REGION Network 7: UN - Hold Command
   RUNG wire#powerrail
      Contact( "UN".PackML_Sts_Alarm.cmd_Hold )
      Contact( "UN".PackML_Sts_Alarm.moduleActive )
      wire#w1
      Coil( "UN".PackML_Sts.cmd_Hold )
   END_RUNG
   RUNG wire#powerrail
      Contact( "EM00".PackML_Sts.Unit.cmd_Hold )
      Contact( "EM00".PackML_Sts.Unit.moduleActive )
   END_RUNG wire#w1
   RUNG wire#powerrail
      Contact( "EM01".PackML_Sts.Unit.cmd_Hold )
      Contact( "EM01".PackML_Sts.Unit.moduleActive )
   END_RUNG wire#w1
   RUNG wire#powerrail
      Contact( "EM02".PackML_Sts.Unit.cmd_Hold )
      Contact( "EM02".PackML_Sts.Unit.moduleActive )
   END_RUNG wire#w1
   // the same network as SCL:
   "UN".PackML_Sts.cmd_Hold := ("UN".PackML_Sts_Alarm.cmd_Hold AND "UN".PackML_Sts_Alarm.moduleActive) OR ("EM00".PackML_Sts.Unit.cmd_Hold AND "EM00".PackML_Sts.Unit.moduleActive) OR ("EM01".PackML_Sts.Unit.cmd_Hold AND "EM01".PackML_Sts.Unit.moduleActive) OR ("EM02".PackML_Sts.Unit.cmd_Hold AND "EM02".PackML_Sts.Unit.moduleActive);
END_REGION

REGION Network 8: UN - Holding State Complete
   RUNG wire#powerrail
      Contact( "UN".PackML_Sts_Alarm.sts_Holding_SC )
      wire#w1
      Contact( "EM00".PackML_Sts.Unit.sts_Holding_SC )
      wire#w2
      Contact( "EM01".PackML_Sts.Unit.sts_Holding_SC )
      wire#w3
      Contact( "EM02".PackML_Sts.Unit.sts_Holding_SC )
      wire#w4
      Coil( "UN".PackML_Sts.sts_Holding_SC )
   END_RUNG
   RUNG wire#powerrail
      I_Contact( "UN".PackML_Sts_Alarm.moduleActive )
   END_RUNG wire#w1
   RUNG wire#w1
      I_Contact( "EM00".PackML_Sts.Unit.moduleActive )
   END_RUNG wire#w2
   RUNG wire#w2
      I_Contact( "EM01".PackML_Sts.Unit.moduleActive )
   END_RUNG wire#w3
   RUNG wire#w3
      I_Contact( "EM02".PackML_Sts.Unit.moduleActive )
   END_RUNG wire#w4
   // the same network as SCL:
   "UN".PackML_Sts.sts_Holding_SC := ("UN".PackML_Sts_Alarm.sts_Holding_SC OR NOT "UN".PackML_Sts_Alarm.moduleActive) AND ("EM00".PackML_Sts.Unit.sts_Holding_SC OR NOT "EM00".PackML_Sts.Unit.moduleActive) AND ("EM01".PackML_Sts.Unit.sts_Holding_SC OR NOT "EM01".PackML_Sts.Unit.moduleActive) AND ("EM02".PackML_Sts.Unit.sts_Holding_SC OR NOT "EM02".PackML_Sts.Unit.moduleActive);
END_REGION

REGION Network 9: UN - UnHold Command
   RUNG wire#powerrail
      Contact( "UN".PackML_Sts_Alarm.cmd_UnHold )
      wire#w1
      Contact( "EM00".PackML_Sts.Unit.cmd_UnHold )
      wire#w2
      Contact( "EM01".PackML_Sts.Unit.cmd_UnHold )
      wire#w3
      Contact( "EM02".PackML_Sts.Unit.cmd_UnHold )
      wire#w4
      Coil( "UN".PackML_Sts.cmd_UnHold )
   END_RUNG
   RUNG wire#powerrail
      I_Contact( "UN".PackML_Sts_Alarm.moduleActive )
   END_RUNG wire#w1
   RUNG wire#w1
      I_Contact( "EM00".PackML_Sts.Unit.moduleActive )
   END_RUNG wire#w2
   RUNG wire#w2
      I_Contact( "EM01".PackML_Sts.Unit.moduleActive )
   END_RUNG wire#w3
   RUNG wire#w3
      I_Contact( "EM02".PackML_Sts.Unit.moduleActive )
   END_RUNG wire#w4
   // the same network as SCL:
   "UN".PackML_Sts.cmd_UnHold := ("UN".PackML_Sts_Alarm.cmd_UnHold OR NOT "UN".PackML_Sts_Alarm.moduleActive) AND ("EM00".PackML_Sts.Unit.cmd_UnHold OR NOT "EM00".PackML_Sts.Unit.moduleActive) AND ("EM01".PackML_Sts.Unit.cmd_UnHold OR NOT "EM01".PackML_Sts.Unit.moduleActive) AND ("EM02".PackML_Sts.Unit.cmd_UnHold OR NOT "EM02".PackML_Sts.Unit.moduleActive);
END_REGION

REGION Network 10: UN - UnHolding State Complete
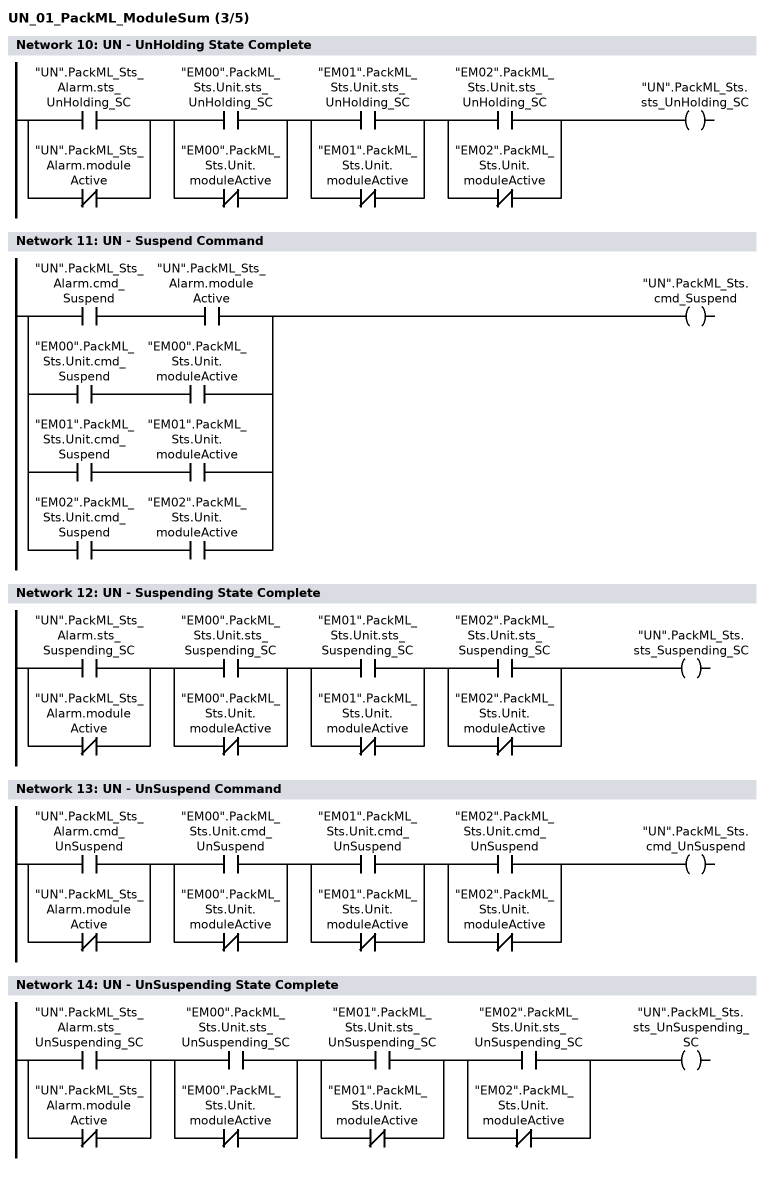
   RUNG wire#powerrail
      Contact( "UN".PackML_Sts_Alarm.sts_UnHolding_SC )
      wire#w1
      Contact( "EM00".PackML_Sts.Unit.sts_UnHolding_SC )
      wire#w2
      Contact( "EM01".PackML_Sts.Unit.sts_UnHolding_SC )
      wire#w3
      Contact( "EM02".PackML_Sts.Unit.sts_UnHolding_SC )
      wire#w4
      Coil( "UN".PackML_Sts.sts_UnHolding_SC )
   END_RUNG
   RUNG wire#powerrail
      I_Contact( "UN".PackML_Sts_Alarm.moduleActive )
   END_RUNG wire#w1
   RUNG wire#w1
      I_Contact( "EM00".PackML_Sts.Unit.moduleActive )
   END_RUNG wire#w2
   RUNG wire#w2
      I_Contact( "EM01".PackML_Sts.Unit.moduleActive )
   END_RUNG wire#w3
   RUNG wire#w3
      I_Contact( "EM02".PackML_Sts.Unit.moduleActive )
   END_RUNG wire#w4
   // the same network as SCL:
   "UN".PackML_Sts.sts_UnHolding_SC := ("UN".PackML_Sts_Alarm.sts_UnHolding_SC OR NOT "UN".PackML_Sts_Alarm.moduleActive) AND ("EM00".PackML_Sts.Unit.sts_UnHolding_SC OR NOT "EM00".PackML_Sts.Unit.moduleActive) AND ("EM01".PackML_Sts.Unit.sts_UnHolding_SC OR NOT "EM01".PackML_Sts.Unit.moduleActive) AND ("EM02".PackML_Sts.Unit.sts_UnHolding_SC OR NOT "EM02".PackML_Sts.Unit.moduleActive);
END_REGION

REGION Network 11: UN - Suspend Command
   RUNG wire#powerrail
      Contact( "UN".PackML_Sts_Alarm.cmd_Suspend )
      Contact( "UN".PackML_Sts_Alarm.moduleActive )
      wire#w1
      Coil( "UN".PackML_Sts.cmd_Suspend )
   END_RUNG
   RUNG wire#powerrail
      Contact( "EM00".PackML_Sts.Unit.cmd_Suspend )
      Contact( "EM00".PackML_Sts.Unit.moduleActive )
   END_RUNG wire#w1
   RUNG wire#powerrail
      Contact( "EM01".PackML_Sts.Unit.cmd_Suspend )
      Contact( "EM01".PackML_Sts.Unit.moduleActive )
   END_RUNG wire#w1
   RUNG wire#powerrail
      Contact( "EM02".PackML_Sts.Unit.cmd_Suspend )
      Contact( "EM02".PackML_Sts.Unit.moduleActive )
   END_RUNG wire#w1
   // the same network as SCL:
   "UN".PackML_Sts.cmd_Suspend := ("UN".PackML_Sts_Alarm.cmd_Suspend AND "UN".PackML_Sts_Alarm.moduleActive) OR ("EM00".PackML_Sts.Unit.cmd_Suspend AND "EM00".PackML_Sts.Unit.moduleActive) OR ("EM01".PackML_Sts.Unit.cmd_Suspend AND "EM01".PackML_Sts.Unit.moduleActive) OR ("EM02".PackML_Sts.Unit.cmd_Suspend AND "EM02".PackML_Sts.Unit.moduleActive);
END_REGION

REGION Network 12: UN - Suspending State Complete
   RUNG wire#powerrail
      Contact( "UN".PackML_Sts_Alarm.sts_Suspending_SC )
      wire#w1
      Contact( "EM00".PackML_Sts.Unit.sts_Suspending_SC )
      wire#w2
      Contact( "EM01".PackML_Sts.Unit.sts_Suspending_SC )
      wire#w3
      Contact( "EM02".PackML_Sts.Unit.sts_Suspending_SC )
      wire#w4
      Coil( "UN".PackML_Sts.sts_Suspending_SC )
   END_RUNG
   RUNG wire#powerrail
      I_Contact( "UN".PackML_Sts_Alarm.moduleActive )
   END_RUNG wire#w1
   RUNG wire#w1
      I_Contact( "EM00".PackML_Sts.Unit.moduleActive )
   END_RUNG wire#w2
   RUNG wire#w2
      I_Contact( "EM01".PackML_Sts.Unit.moduleActive )
   END_RUNG wire#w3
   RUNG wire#w3
      I_Contact( "EM02".PackML_Sts.Unit.moduleActive )
   END_RUNG wire#w4
   // the same network as SCL:
   "UN".PackML_Sts.sts_Suspending_SC := ("UN".PackML_Sts_Alarm.sts_Suspending_SC OR NOT "UN".PackML_Sts_Alarm.moduleActive) AND ("EM00".PackML_Sts.Unit.sts_Suspending_SC OR NOT "EM00".PackML_Sts.Unit.moduleActive) AND ("EM01".PackML_Sts.Unit.sts_Suspending_SC OR NOT "EM01".PackML_Sts.Unit.moduleActive) AND ("EM02".PackML_Sts.Unit.sts_Suspending_SC OR NOT "EM02".PackML_Sts.Unit.moduleActive);
END_REGION

REGION Network 13: UN - UnSuspend Command
   RUNG wire#powerrail
      Contact( "UN".PackML_Sts_Alarm.cmd_UnSuspend )
      wire#w1
      Contact( "EM00".PackML_Sts.Unit.cmd_UnSuspend )
      wire#w2
      Contact( "EM01".PackML_Sts.Unit.cmd_UnSuspend )
      wire#w3
      Contact( "EM02".PackML_Sts.Unit.cmd_UnSuspend )
      wire#w4
      Coil( "UN".PackML_Sts.cmd_UnSuspend )
   END_RUNG
   RUNG wire#powerrail
      I_Contact( "UN".PackML_Sts_Alarm.moduleActive )
   END_RUNG wire#w1
   RUNG wire#w1
      I_Contact( "EM00".PackML_Sts.Unit.moduleActive )
   END_RUNG wire#w2
   RUNG wire#w2
      I_Contact( "EM01".PackML_Sts.Unit.moduleActive )
   END_RUNG wire#w3
   RUNG wire#w3
      I_Contact( "EM02".PackML_Sts.Unit.moduleActive )
   END_RUNG wire#w4
   // the same network as SCL:
   "UN".PackML_Sts.cmd_UnSuspend := ("UN".PackML_Sts_Alarm.cmd_UnSuspend OR NOT "UN".PackML_Sts_Alarm.moduleActive) AND ("EM00".PackML_Sts.Unit.cmd_UnSuspend OR NOT "EM00".PackML_Sts.Unit.moduleActive) AND ("EM01".PackML_Sts.Unit.cmd_UnSuspend OR NOT "EM01".PackML_Sts.Unit.moduleActive) AND ("EM02".PackML_Sts.Unit.cmd_UnSuspend OR NOT "EM02".PackML_Sts.Unit.moduleActive);
END_REGION

REGION Network 14: UN - UnSuspending State Complete
   RUNG wire#powerrail
      Contact( "UN".PackML_Sts_Alarm.sts_UnSuspending_SC )
      wire#w1
      Contact( "EM00".PackML_Sts.Unit.sts_UnSuspending_SC )
      wire#w2
      Contact( "EM01".PackML_Sts.Unit.sts_UnSuspending_SC )
      wire#w3
      Contact( "EM02".PackML_Sts.Unit.sts_UnSuspending_SC )
      wire#w4
      Coil( "UN".PackML_Sts.sts_UnSuspending_SC )
   END_RUNG
   RUNG wire#powerrail
      I_Contact( "UN".PackML_Sts_Alarm.moduleActive )
   END_RUNG wire#w1
   RUNG wire#w1
      I_Contact( "EM00".PackML_Sts.Unit.moduleActive )
   END_RUNG wire#w2
   RUNG wire#w2
      I_Contact( "EM01".PackML_Sts.Unit.moduleActive )
   END_RUNG wire#w3
   RUNG wire#w3
      I_Contact( "EM02".PackML_Sts.Unit.moduleActive )
   END_RUNG wire#w4
   // the same network as SCL:
   "UN".PackML_Sts.sts_UnSuspending_SC := ("UN".PackML_Sts_Alarm.sts_UnSuspending_SC OR NOT "UN".PackML_Sts_Alarm.moduleActive) AND ("EM00".PackML_Sts.Unit.sts_UnSuspending_SC OR NOT "EM00".PackML_Sts.Unit.moduleActive) AND ("EM01".PackML_Sts.Unit.sts_UnSuspending_SC OR NOT "EM01".PackML_Sts.Unit.moduleActive) AND ("EM02".PackML_Sts.Unit.sts_UnSuspending_SC OR NOT "EM02".PackML_Sts.Unit.moduleActive);
END_REGION

REGION Network 15: UN - Abort Command
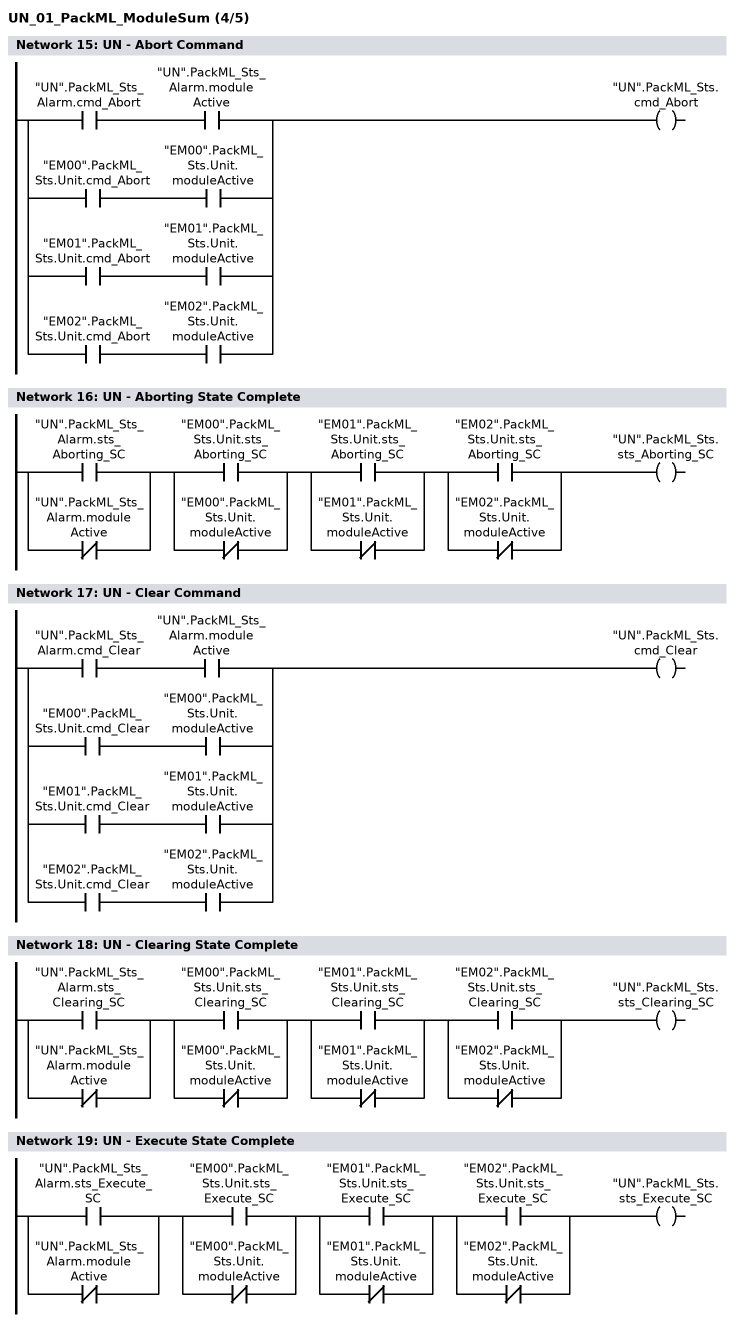
   RUNG wire#powerrail
      Contact( "UN".PackML_Sts_Alarm.cmd_Abort )
      Contact( "UN".PackML_Sts_Alarm.moduleActive )
      wire#w1
      Coil( "UN".PackML_Sts.cmd_Abort )
   END_RUNG
   RUNG wire#powerrail
      Contact( "EM00".PackML_Sts.Unit.cmd_Abort )
      Contact( "EM00".PackML_Sts.Unit.moduleActive )
   END_RUNG wire#w1
   RUNG wire#powerrail
      Contact( "EM01".PackML_Sts.Unit.cmd_Abort )
      Contact( "EM01".PackML_Sts.Unit.moduleActive )
   END_RUNG wire#w1
   RUNG wire#powerrail
      Contact( "EM02".PackML_Sts.Unit.cmd_Abort )
      Contact( "EM02".PackML_Sts.Unit.moduleActive )
   END_RUNG wire#w1
   // the same network as SCL:
   "UN".PackML_Sts.cmd_Abort := ("UN".PackML_Sts_Alarm.cmd_Abort AND "UN".PackML_Sts_Alarm.moduleActive) OR ("EM00".PackML_Sts.Unit.cmd_Abort AND "EM00".PackML_Sts.Unit.moduleActive) OR ("EM01".PackML_Sts.Unit.cmd_Abort AND "EM01".PackML_Sts.Unit.moduleActive) OR ("EM02".PackML_Sts.Unit.cmd_Abort AND "EM02".PackML_Sts.Unit.moduleActive);
END_REGION

REGION Network 16: UN - Aborting State Complete
   RUNG wire#powerrail
      Contact( "UN".PackML_Sts_Alarm.sts_Aborting_SC )
      wire#w1
      Contact( "EM00".PackML_Sts.Unit.sts_Aborting_SC )
      wire#w2
      Contact( "EM01".PackML_Sts.Unit.sts_Aborting_SC )
      wire#w3
      Contact( "EM02".PackML_Sts.Unit.sts_Aborting_SC )
      wire#w4
      Coil( "UN".PackML_Sts.sts_Aborting_SC )
   END_RUNG
   RUNG wire#powerrail
      I_Contact( "UN".PackML_Sts_Alarm.moduleActive )
   END_RUNG wire#w1
   RUNG wire#w1
      I_Contact( "EM00".PackML_Sts.Unit.moduleActive )
   END_RUNG wire#w2
   RUNG wire#w2
      I_Contact( "EM01".PackML_Sts.Unit.moduleActive )
   END_RUNG wire#w3
   RUNG wire#w3
      I_Contact( "EM02".PackML_Sts.Unit.moduleActive )
   END_RUNG wire#w4
   // the same network as SCL:
   "UN".PackML_Sts.sts_Aborting_SC := ("UN".PackML_Sts_Alarm.sts_Aborting_SC OR NOT "UN".PackML_Sts_Alarm.moduleActive) AND ("EM00".PackML_Sts.Unit.sts_Aborting_SC OR NOT "EM00".PackML_Sts.Unit.moduleActive) AND ("EM01".PackML_Sts.Unit.sts_Aborting_SC OR NOT "EM01".PackML_Sts.Unit.moduleActive) AND ("EM02".PackML_Sts.Unit.sts_Aborting_SC OR NOT "EM02".PackML_Sts.Unit.moduleActive);
END_REGION

REGION Network 17: UN - Clear Command
   RUNG wire#powerrail
      Contact( "UN".PackML_Sts_Alarm.cmd_Clear )
      Contact( "UN".PackML_Sts_Alarm.moduleActive )
      wire#w1
      Coil( "UN".PackML_Sts.cmd_Clear )
   END_RUNG
   RUNG wire#powerrail
      Contact( "EM00".PackML_Sts.Unit.cmd_Clear )
      Contact( "EM00".PackML_Sts.Unit.moduleActive )
   END_RUNG wire#w1
   RUNG wire#powerrail
      Contact( "EM01".PackML_Sts.Unit.cmd_Clear )
      Contact( "EM01".PackML_Sts.Unit.moduleActive )
   END_RUNG wire#w1
   RUNG wire#powerrail
      Contact( "EM02".PackML_Sts.Unit.cmd_Clear )
      Contact( "EM02".PackML_Sts.Unit.moduleActive )
   END_RUNG wire#w1
   // the same network as SCL:
   "UN".PackML_Sts.cmd_Clear := ("UN".PackML_Sts_Alarm.cmd_Clear AND "UN".PackML_Sts_Alarm.moduleActive) OR ("EM00".PackML_Sts.Unit.cmd_Clear AND "EM00".PackML_Sts.Unit.moduleActive) OR ("EM01".PackML_Sts.Unit.cmd_Clear AND "EM01".PackML_Sts.Unit.moduleActive) OR ("EM02".PackML_Sts.Unit.cmd_Clear AND "EM02".PackML_Sts.Unit.moduleActive);
END_REGION

REGION Network 18: UN - Clearing State Complete
   RUNG wire#powerrail
      Contact( "UN".PackML_Sts_Alarm.sts_Clearing_SC )
      wire#w1
      Contact( "EM00".PackML_Sts.Unit.sts_Clearing_SC )
      wire#w2
      Contact( "EM01".PackML_Sts.Unit.sts_Clearing_SC )
      wire#w3
      Contact( "EM02".PackML_Sts.Unit.sts_Clearing_SC )
      wire#w4
      Coil( "UN".PackML_Sts.sts_Clearing_SC )
   END_RUNG
   RUNG wire#powerrail
      I_Contact( "UN".PackML_Sts_Alarm.moduleActive )
   END_RUNG wire#w1
   RUNG wire#w1
      I_Contact( "EM00".PackML_Sts.Unit.moduleActive )
   END_RUNG wire#w2
   RUNG wire#w2
      I_Contact( "EM01".PackML_Sts.Unit.moduleActive )
   END_RUNG wire#w3
   RUNG wire#w3
      I_Contact( "EM02".PackML_Sts.Unit.moduleActive )
   END_RUNG wire#w4
   // the same network as SCL:
   "UN".PackML_Sts.sts_Clearing_SC := ("UN".PackML_Sts_Alarm.sts_Clearing_SC OR NOT "UN".PackML_Sts_Alarm.moduleActive) AND ("EM00".PackML_Sts.Unit.sts_Clearing_SC OR NOT "EM00".PackML_Sts.Unit.moduleActive) AND ("EM01".PackML_Sts.Unit.sts_Clearing_SC OR NOT "EM01".PackML_Sts.Unit.moduleActive) AND ("EM02".PackML_Sts.Unit.sts_Clearing_SC OR NOT "EM02".PackML_Sts.Unit.moduleActive);
END_REGION

REGION Network 19: UN - Execute State Complete
   RUNG wire#powerrail
      Contact( "UN".PackML_Sts_Alarm.sts_Execute_SC )
      wire#w1
      Contact( "EM00".PackML_Sts.Unit.sts_Execute_SC )
      wire#w2
      Contact( "EM01".PackML_Sts.Unit.sts_Execute_SC )
      wire#w3
      Contact( "EM02".PackML_Sts.Unit.sts_Execute_SC )
      wire#w4
      Coil( "UN".PackML_Sts.sts_Execute_SC )
   END_RUNG
   RUNG wire#powerrail
      I_Contact( "UN".PackML_Sts_Alarm.moduleActive )
   END_RUNG wire#w1
   RUNG wire#w1
      I_Contact( "EM00".PackML_Sts.Unit.moduleActive )
   END_RUNG wire#w2
   RUNG wire#w2
      I_Contact( "EM01".PackML_Sts.Unit.moduleActive )
   END_RUNG wire#w3
   RUNG wire#w3
      I_Contact( "EM02".PackML_Sts.Unit.moduleActive )
   END_RUNG wire#w4
   // the same network as SCL:
   "UN".PackML_Sts.sts_Execute_SC := ("UN".PackML_Sts_Alarm.sts_Execute_SC OR NOT "UN".PackML_Sts_Alarm.moduleActive) AND ("EM00".PackML_Sts.Unit.sts_Execute_SC OR NOT "EM00".PackML_Sts.Unit.moduleActive) AND ("EM01".PackML_Sts.Unit.sts_Execute_SC OR NOT "EM01".PackML_Sts.Unit.moduleActive) AND ("EM02".PackML_Sts.Unit.sts_Execute_SC OR NOT "EM02".PackML_Sts.Unit.moduleActive);
END_REGION

REGION Network 20: UN - Completing State Complete
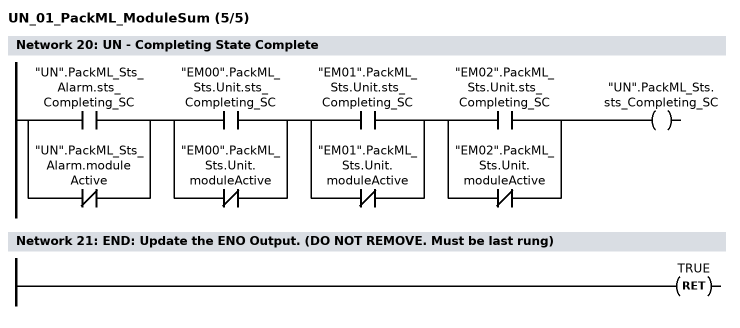
   RUNG wire#powerrail
      Contact( "UN".PackML_Sts_Alarm.sts_Completing_SC )
      wire#w1
      Contact( "EM00".PackML_Sts.Unit.sts_Completing_SC )
      wire#w2
      Contact( "EM01".PackML_Sts.Unit.sts_Completing_SC )
      wire#w3
      Contact( "EM02".PackML_Sts.Unit.sts_Completing_SC )
      wire#w4
      Coil( "UN".PackML_Sts.sts_Completing_SC )
   END_RUNG
   RUNG wire#powerrail
      I_Contact( "UN".PackML_Sts_Alarm.moduleActive )
   END_RUNG wire#w1
   RUNG wire#w1
      I_Contact( "EM00".PackML_Sts.Unit.moduleActive )
   END_RUNG wire#w2
   RUNG wire#w2
      I_Contact( "EM01".PackML_Sts.Unit.moduleActive )
   END_RUNG wire#w3
   RUNG wire#w3
      I_Contact( "EM02".PackML_Sts.Unit.moduleActive )
   END_RUNG wire#w4
   // the same network as SCL:
   "UN".PackML_Sts.sts_Completing_SC := ("UN".PackML_Sts_Alarm.sts_Completing_SC OR NOT "UN".PackML_Sts_Alarm.moduleActive) AND ("EM00".PackML_Sts.Unit.sts_Completing_SC OR NOT "EM00".PackML_Sts.Unit.moduleActive) AND ("EM01".PackML_Sts.Unit.sts_Completing_SC OR NOT "EM01".PackML_Sts.Unit.moduleActive) AND ("EM02".PackML_Sts.Unit.sts_Completing_SC OR NOT "EM02".PackML_Sts.Unit.moduleActive);
END_REGION

REGION Network 21: END: Update the ENO Output. (DO NOT REMOVE. Must be last rung)
   RUNG wire#powerrail
      ReturnCoil( TRUE )
   END_RUNG
   // the same network as SCL:
   ENO := TRUE;
   RETURN;
END_REGION
END_FUNCTION_BLOCK

FUNCTION_BLOCK "UN_02_PackML"   // FB31622, LAD
TITLE = UN_02_PackML
{ S7_Optimized_Access := 'TRUE' }
AUTHOR : tech.team.motioncontrol@siemens.com
FAMILY : CPG
VERSION : 1.0
// Support: tech.team.motioncontrol@siemens.com
// Fax: +49 (0) 9131/98-1297
   VAR
      statLanguageSelectedOld : Int := -1;
      statPackML_CMD_SC : Bool;
      instUnitModeStateManager : "LPMLV30_UnitModeStateManager";
      instUnitModeStateTimes : "LPMLV30_UnitModeStateTimes";
      statRemoteCommand_ModeChangeRequest : Struct
         Production : Bool;   // Request to goto mode - PRODUCTION (mode #1)
         Maintenance : Bool;   // Request to goto mode - MAINTENANCE (mode #2)
         Manual : Bool;   // Request to goto mode - MANUAL (mode #3)
         UserMode01 : Bool;   // Request to goto mode - USER MODE 01 (mode #4)
         UserMode02 : Bool;   // Request to goto mode - USER MODE 02 (mode #5)
         UserMode03 : Bool;   // Request to goto mode - USER MODE 03 (mode #6)
         UserMode04 : Bool;   // Request to goto mode - USER MODE 04 (mode #7)
         UserMode05 : Bool;   // Request to goto mode - USER MODE 05 (mode #8)
         UserMode06 : Bool;   // Request to goto mode - USER MODE 06 (mode #9)
         UserMode07 : Bool;   // Request to goto mode - USER MODE 07 (mode #10)
         UserMode08 : Bool;   // Request to goto mode - USER MODE 08 (mode #11)
      END_STRUCT;
      TPResettingDelay : TP_TIME;
      TPClearingDelay : TP_TIME;
   END_VAR
   VAR_TEMP
      tempDiagnosticsBufferIndexForHMI : Int;   // Temporary integer for PackML HMI diagnostics
   END_VAR
   VAR_TEMP   // added for the SCL form of the ladder/FBD networks
      _w1 : Bool;
   END_VAR
BEGIN

REGION Network 1: PackML ModeManager & State Model - Reset command
   // Reset Command:
   // If the machine is stopped and there are no faults (no stop or abort commands), 
   // then automatically reset and move the machine to idle.  This is common when all 
   // the faults are cleared in the Clearing state and the machine moves to the 
   // Stopped state with no more faults.
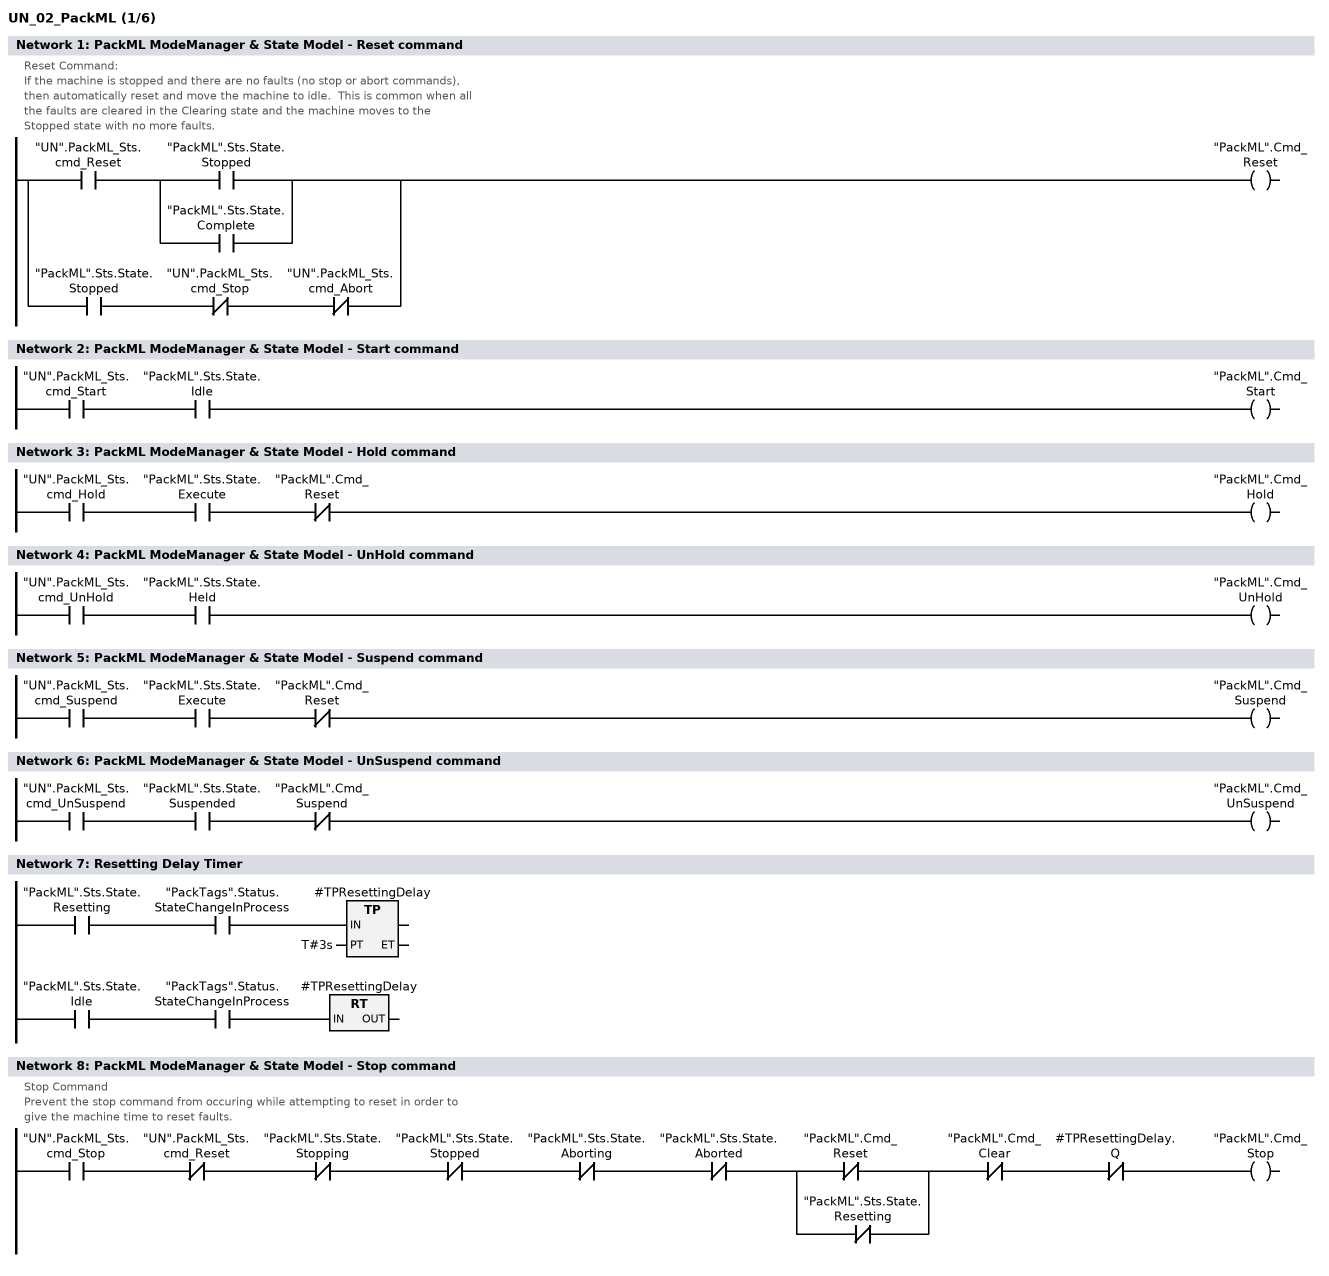
   RUNG wire#powerrail
      Contact( "UN".PackML_Sts.cmd_Reset )
      wire#w1
      Contact( "PackML".Sts.State.Stopped )
      wire#w2
      Coil( "PackML".Cmd_Reset )
   END_RUNG
   RUNG wire#w1
      Contact( "PackML".Sts.State.Complete )
   END_RUNG wire#w2
   RUNG wire#powerrail
      Contact( "PackML".Sts.State.Stopped )
      I_Contact( "UN".PackML_Sts.cmd_Stop )
      I_Contact( "UN".PackML_Sts.cmd_Abort )
   END_RUNG wire#w2
   // the same network as SCL:
   "PackML".Cmd_Reset := ("UN".PackML_Sts.cmd_Reset AND ("PackML".Sts.State.Stopped OR "PackML".Sts.State.Complete)) OR ("PackML".Sts.State.Stopped AND NOT "UN".PackML_Sts.cmd_Stop AND NOT "UN".PackML_Sts.cmd_Abort);
END_REGION

REGION Network 2: PackML ModeManager & State Model - Start command
   RUNG wire#powerrail
      Contact( "UN".PackML_Sts.cmd_Start )
      Contact( "PackML".Sts.State.Idle )
      Coil( "PackML".Cmd_Start )
   END_RUNG
   // the same network as SCL:
   "PackML".Cmd_Start := "UN".PackML_Sts.cmd_Start AND "PackML".Sts.State.Idle;
END_REGION

REGION Network 3: PackML ModeManager & State Model - Hold command
   RUNG wire#powerrail
      Contact( "UN".PackML_Sts.cmd_Hold )
      Contact( "PackML".Sts.State.Execute )
      I_Contact( "PackML".Cmd_Reset )
      Coil( "PackML".Cmd_Hold )
   END_RUNG
   // the same network as SCL:
   "PackML".Cmd_Hold := "UN".PackML_Sts.cmd_Hold AND "PackML".Sts.State.Execute AND NOT "PackML".Cmd_Reset;
END_REGION

REGION Network 4: PackML ModeManager & State Model - UnHold command
   RUNG wire#powerrail
      Contact( "UN".PackML_Sts.cmd_UnHold )
      Contact( "PackML".Sts.State.Held )
      Coil( "PackML".Cmd_UnHold )
   END_RUNG
   // the same network as SCL:
   "PackML".Cmd_UnHold := "UN".PackML_Sts.cmd_UnHold AND "PackML".Sts.State.Held;
END_REGION

REGION Network 5: PackML ModeManager & State Model - Suspend command
   RUNG wire#powerrail
      Contact( "UN".PackML_Sts.cmd_Suspend )
      Contact( "PackML".Sts.State.Execute )
      I_Contact( "PackML".Cmd_Reset )
      Coil( "PackML".Cmd_Suspend )
   END_RUNG
   // the same network as SCL:
   "PackML".Cmd_Suspend := "UN".PackML_Sts.cmd_Suspend AND "PackML".Sts.State.Execute AND NOT "PackML".Cmd_Reset;
END_REGION

REGION Network 6: PackML ModeManager & State Model - UnSuspend command
   RUNG wire#powerrail
      Contact( "UN".PackML_Sts.cmd_UnSuspend )
      Contact( "PackML".Sts.State.Suspended )
      I_Contact( "PackML".Cmd_Suspend )
      Coil( "PackML".Cmd_UnSuspend )
   END_RUNG
   // the same network as SCL:
   "PackML".Cmd_UnSuspend := "UN".PackML_Sts.cmd_UnSuspend AND "PackML".Sts.State.Suspended AND NOT "PackML".Cmd_Suspend;
END_REGION

REGION Network 7: Resetting Delay Timer
   #TPResettingDelay(IN := "PackML".Sts.State.Resetting AND "PackTags".Status.StateChangeInProcess, PT := T#3s);   // TP
   IF "PackML".Sts.State.Idle AND "PackTags".Status.StateChangeInProcess THEN
       RESET_TIMER(#TPResettingDelay);
   END_IF;
END_REGION

REGION Network 8: PackML ModeManager & State Model - Stop command
   // Stop Command
   // Prevent the stop command from occuring while attempting to reset in order to 
   // give the machine time to reset faults.
   RUNG wire#powerrail
      Contact( "UN".PackML_Sts.cmd_Stop )
      I_Contact( "UN".PackML_Sts.cmd_Reset )
      I_Contact( "PackML".Sts.State.Stopping )
      I_Contact( "PackML".Sts.State.Stopped )
      I_Contact( "PackML".Sts.State.Aborting )
      I_Contact( "PackML".Sts.State.Aborted )
      wire#w1
      I_Contact( "PackML".Cmd_Reset )
      wire#w2
      I_Contact( "PackML".Cmd_Clear )
      I_Contact( #TPResettingDelay.Q )
      Coil( "PackML".Cmd_Stop )
   END_RUNG
   RUNG wire#w1
      I_Contact( "PackML".Sts.State.Resetting )
   END_RUNG wire#w2
   // the same network as SCL:
   "PackML".Cmd_Stop := "UN".PackML_Sts.cmd_Stop AND NOT "UN".PackML_Sts.cmd_Reset AND NOT "PackML".Sts.State.Stopping AND NOT "PackML".Sts.State.Stopped AND NOT "PackML".Sts.State.Aborting AND NOT "PackML".Sts.State.Aborted AND (NOT "PackML".Cmd_Reset OR NOT "PackML".Sts.State.Resetting) AND NOT "PackML".Cmd_Clear AND NOT #TPResettingDelay.Q;
END_REGION

REGION Network 9: Clearing Delay Timer
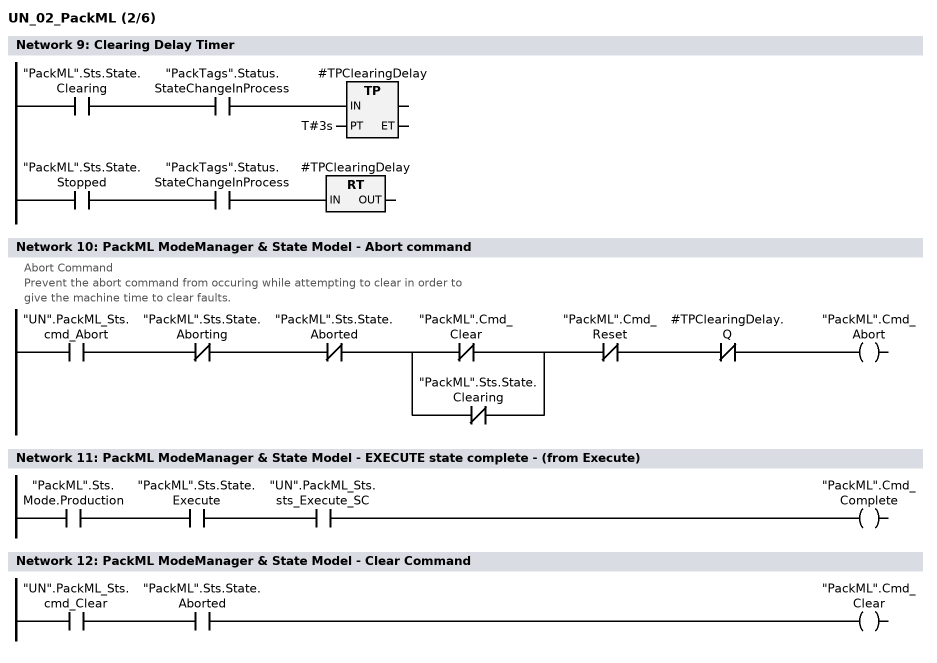
   #TPClearingDelay(IN := "PackML".Sts.State.Clearing AND "PackTags".Status.StateChangeInProcess, PT := T#3s);   // TP
   IF "PackML".Sts.State.Stopped AND "PackTags".Status.StateChangeInProcess THEN
       RESET_TIMER(#TPClearingDelay);
   END_IF;
END_REGION

REGION Network 10: PackML ModeManager & State Model - Abort command
   // Abort Command
   // Prevent the abort command from occuring while attempting to clear in order to 
   // give the machine time to clear faults.
   RUNG wire#powerrail
      Contact( "UN".PackML_Sts.cmd_Abort )
      I_Contact( "PackML".Sts.State.Aborting )
      I_Contact( "PackML".Sts.State.Aborted )
      wire#w1
      I_Contact( "PackML".Cmd_Clear )
      wire#w2
      I_Contact( "PackML".Cmd_Reset )
      I_Contact( #TPClearingDelay.Q )
      Coil( "PackML".Cmd_Abort )
   END_RUNG
   RUNG wire#w1
      I_Contact( "PackML".Sts.State.Clearing )
   END_RUNG wire#w2
   // the same network as SCL:
   "PackML".Cmd_Abort := "UN".PackML_Sts.cmd_Abort AND NOT "PackML".Sts.State.Aborting AND NOT "PackML".Sts.State.Aborted AND (NOT "PackML".Cmd_Clear OR NOT "PackML".Sts.State.Clearing) AND NOT "PackML".Cmd_Reset AND NOT #TPClearingDelay.Q;
END_REGION

REGION Network 11: PackML ModeManager & State Model - EXECUTE state complete - (from Execute)
   RUNG wire#powerrail
      Contact( "PackML".Sts.Mode.Production )
      Contact( "PackML".Sts.State.Execute )
      Contact( "UN".PackML_Sts.sts_Execute_SC )
      Coil( "PackML".Cmd_Complete )
   END_RUNG
   // the same network as SCL:
   "PackML".Cmd_Complete := "PackML".Sts.Mode.Production AND "PackML".Sts.State.Execute AND "UN".PackML_Sts.sts_Execute_SC;
END_REGION

REGION Network 12: PackML ModeManager & State Model - Clear Command
   RUNG wire#powerrail
      Contact( "UN".PackML_Sts.cmd_Clear )
      Contact( "PackML".Sts.State.Aborted )
      Coil( "PackML".Cmd_Clear )
   END_RUNG
   // the same network as SCL:
   "PackML".Cmd_Clear := "UN".PackML_Sts.cmd_Clear AND "PackML".Sts.State.Aborted;
END_REGION

REGION Network 13: External PackML Mode Commands
   // External State Commands are handled in the UN_05_EventControl routine to ensure that the unit machine level alarm manager captures the reason for any machine stoppage.
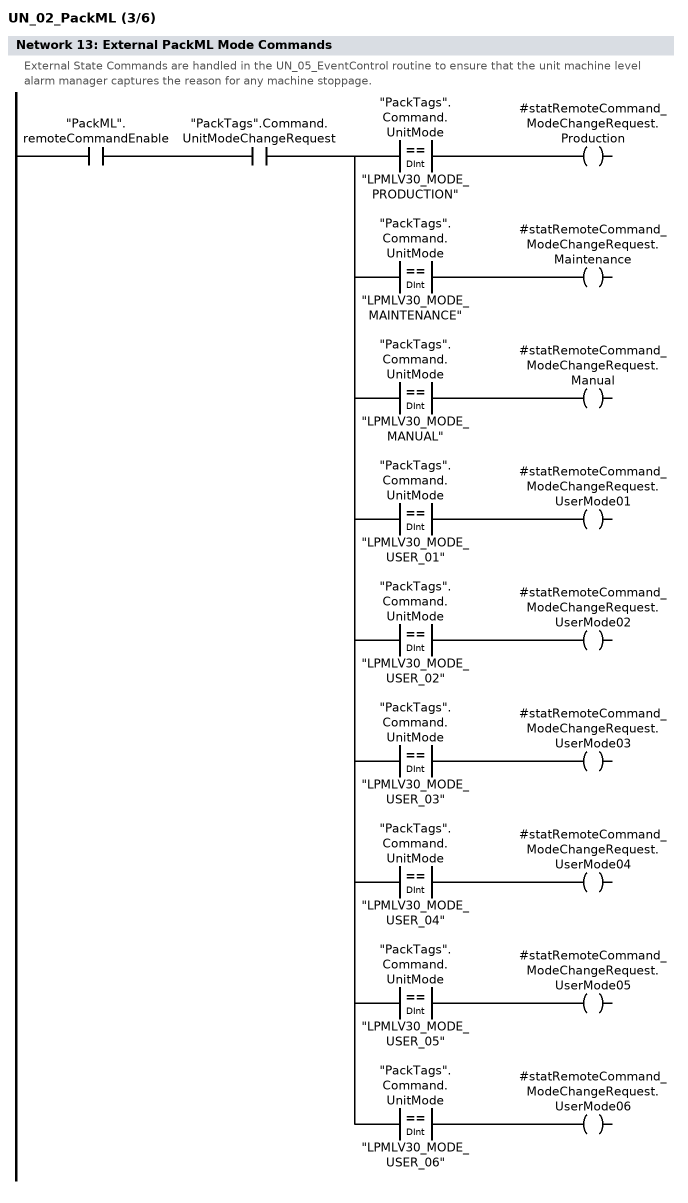
   RUNG wire#powerrail
      Contact( "PackML".remoteCommandEnable )
      Contact( "PackTags".Command.UnitModeChangeRequest )
      wire#w1
      { S7_Templates := "SrcType := DInt" } EQ_Contact(in1 := "PackTags".Command.UnitMode, in2 := "LPMLV30_MODE_PRODUCTION")
      Coil( #statRemoteCommand_ModeChangeRequest.Production )
   END_RUNG
   RUNG wire#w1
      { S7_Templates := "SrcType := DInt" } EQ_Contact(in1 := "PackTags".Command.UnitMode, in2 := "LPMLV30_MODE_MAINTENANCE")
      Coil( #statRemoteCommand_ModeChangeRequest.Maintenance )
   END_RUNG
   RUNG wire#w1
      { S7_Templates := "SrcType := DInt" } EQ_Contact(in1 := "PackTags".Command.UnitMode, in2 := "LPMLV30_MODE_MANUAL")
      Coil( #statRemoteCommand_ModeChangeRequest.Manual )
   END_RUNG
   RUNG wire#w1
      { S7_Templates := "SrcType := DInt" } EQ_Contact(in1 := "PackTags".Command.UnitMode, in2 := "LPMLV30_MODE_USER_01")
      Coil( #statRemoteCommand_ModeChangeRequest.UserMode01 )
   END_RUNG
   RUNG wire#w1
      { S7_Templates := "SrcType := DInt" } EQ_Contact(in1 := "PackTags".Command.UnitMode, in2 := "LPMLV30_MODE_USER_02")
      Coil( #statRemoteCommand_ModeChangeRequest.UserMode02 )
   END_RUNG
   RUNG wire#w1
      { S7_Templates := "SrcType := DInt" } EQ_Contact(in1 := "PackTags".Command.UnitMode, in2 := "LPMLV30_MODE_USER_03")
      Coil( #statRemoteCommand_ModeChangeRequest.UserMode03 )
   END_RUNG
   RUNG wire#w1
      { S7_Templates := "SrcType := DInt" } EQ_Contact(in1 := "PackTags".Command.UnitMode, in2 := "LPMLV30_MODE_USER_04")
      Coil( #statRemoteCommand_ModeChangeRequest.UserMode04 )
   END_RUNG
   RUNG wire#w1
      { S7_Templates := "SrcType := DInt" } EQ_Contact(in1 := "PackTags".Command.UnitMode, in2 := "LPMLV30_MODE_USER_05")
      Coil( #statRemoteCommand_ModeChangeRequest.UserMode05 )
   END_RUNG
   RUNG wire#w1
      { S7_Templates := "SrcType := DInt" } EQ_Contact(in1 := "PackTags".Command.UnitMode, in2 := "LPMLV30_MODE_USER_06")
      Coil( #statRemoteCommand_ModeChangeRequest.UserMode06 )
   END_RUNG
   // the same network as SCL:
   #_w1 := "PackML".remoteCommandEnable AND "PackTags".Command.UnitModeChangeRequest;
   #statRemoteCommand_ModeChangeRequest.Production := #_w1 AND ("PackTags".Command.UnitMode = "LPMLV30_MODE_PRODUCTION");
   #statRemoteCommand_ModeChangeRequest.Maintenance := #_w1 AND ("PackTags".Command.UnitMode = "LPMLV30_MODE_MAINTENANCE");
   #statRemoteCommand_ModeChangeRequest.Manual := #_w1 AND ("PackTags".Command.UnitMode = "LPMLV30_MODE_MANUAL");
   #statRemoteCommand_ModeChangeRequest.UserMode01 := #_w1 AND ("PackTags".Command.UnitMode = "LPMLV30_MODE_USER_01");
   #statRemoteCommand_ModeChangeRequest.UserMode02 := #_w1 AND ("PackTags".Command.UnitMode = "LPMLV30_MODE_USER_02");
   #statRemoteCommand_ModeChangeRequest.UserMode03 := #_w1 AND ("PackTags".Command.UnitMode = "LPMLV30_MODE_USER_03");
   #statRemoteCommand_ModeChangeRequest.UserMode04 := #_w1 AND ("PackTags".Command.UnitMode = "LPMLV30_MODE_USER_04");
   #statRemoteCommand_ModeChangeRequest.UserMode05 := #_w1 AND ("PackTags".Command.UnitMode = "LPMLV30_MODE_USER_05");
   #statRemoteCommand_ModeChangeRequest.UserMode06 := #_w1 AND ("PackTags".Command.UnitMode = "LPMLV30_MODE_USER_06");
END_REGION

REGION Network 14: Call thePackML Mode Manager & State Model FB
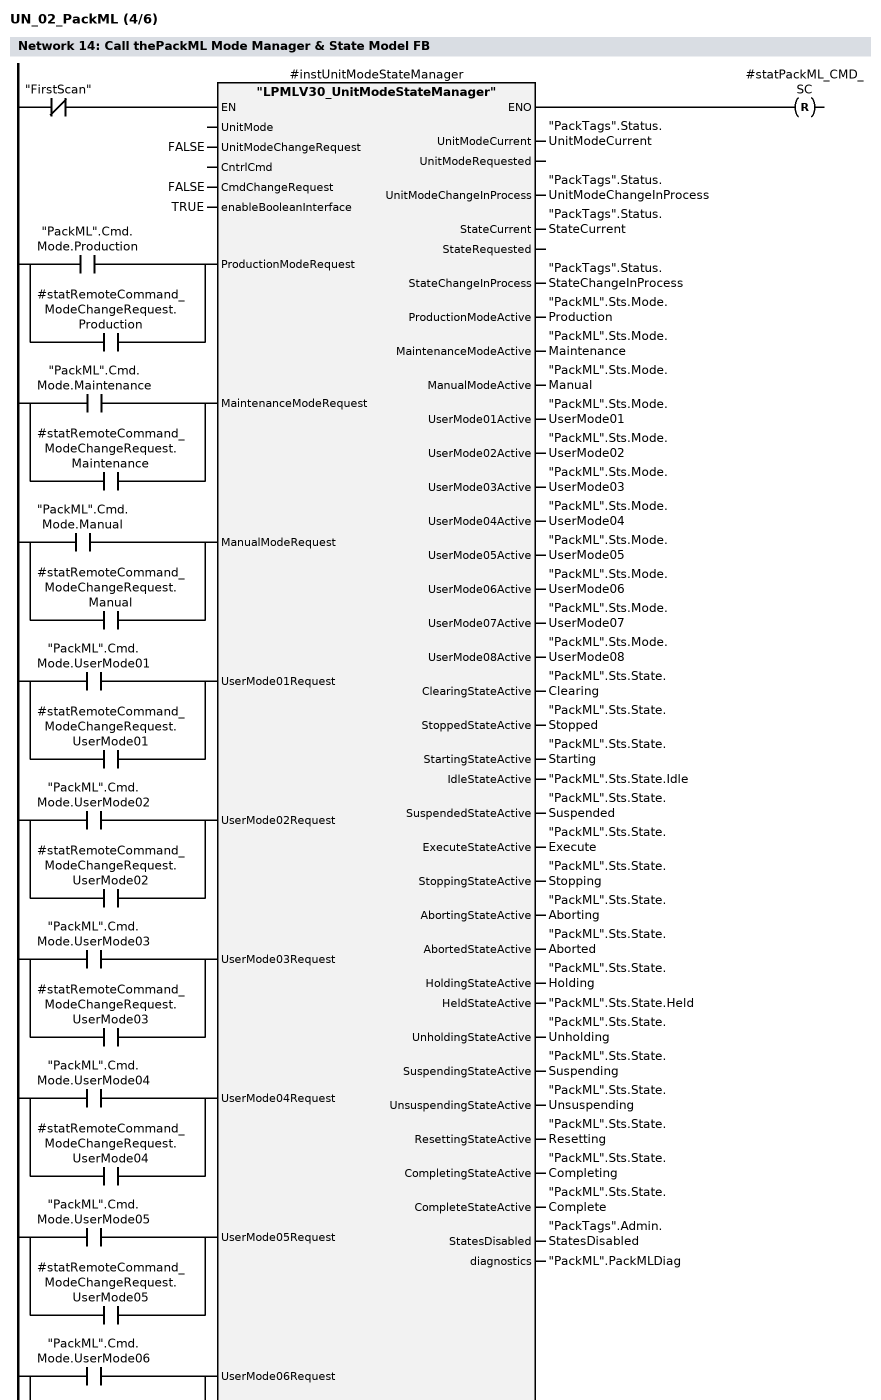